   "煤粉仓温度高报警" AT %Q5.1 : Bool;
   "回转窑助燃罗茨风机启动" AT %Q4.7 : Bool;
   "Q3_7" AT %Q3.7 : Bool;
   "Q3_6" AT %Q3.6 : Bool;
   "Q3_5" AT %Q3.5 : Bool;
   "Q3_4" AT %Q3.4 : Bool;
   "Q3_3" AT %Q3.3 : Bool;
   "Q3_2" AT %Q3.2 : Bool;
   "Q3_1" AT %Q3.1 : Bool;
   "Q3_0" AT %Q3.0 : Bool;
   "Q2_7" AT %Q2.7 : Bool;
   "Q2_6" AT %Q2.6 : Bool;
   "Q2_5" AT %Q2.5 : Bool;
   "Q2_4" AT %Q2.4 : Bool;
   "Q2_3" AT %Q2.3 : Bool;
   "Q2_2" AT %Q2.2 : Bool;
   "Q2_1" AT %Q2.1 : Bool;
   "Q2_0" AT %Q2.0 : Bool;
   "Q1_7" AT %Q1.7 : Bool;
   "Q1_1" AT %Q1.1 : Bool;
   "窑尾罩温度输出" AT %QW286 : Int;
   "PQW278" AT %QW278 : Int;
   "4#回转窑富氧调节阀给定" AT %QW276 : Int;
   "助燃罗茨风机频率给定" AT %QW274 : Int;
   "PQW270" AT %QW270 : Int;
   "PQW268" AT %QW268 : Int;
   "PQW266" AT %QW266 : Int;
   "PQW264" AT %QW264 : Int;
   "PQW262" AT %QW262 : Int;
   "PQW260" AT %QW260 : Int;
   "7#配料皮带启动" AT %Q6.6 : Bool;
   "7#配料流量给定" AT %QW300 : Int;
   "6#配料皮带启动" AT %Q6.5 : Bool;
   "6#配料流量给定" AT %QW298 : Int;
   "5#配料皮带启动" AT %Q6.4 : Bool;
   "5#配料流量给定" AT %QW296 : Int;
   "4#配料皮带启动" AT %Q6.3 : Bool;
   "4#配料流量给定" AT %QW294 : Int;
   "3#配料皮带启动" AT %Q6.2 : Bool;
   "3#配料流量给定" AT %QW292 : Int;
   "2#配料皮带启动" AT %Q6.1 : Bool;
   "2#配料流量给定" AT %QW290 : Int;
   "1#配料皮带启动" AT %Q6.0 : Bool;
   "1#配料流量给定" AT %QW288 : Int;
   "闸阀下限" AT %M80.7 : Bool;
   "闸阀上限" AT %M80.6 : Bool;
   "窑体行程下下限停窑计时" AT %M8.1 : Bool;
   "窑体行程上上限停窑计时" AT %M8.0 : Bool;
   "挡轮油站重故障_BOOL" AT %M10.2 : Bool;
   "回转窑转子秤连锁" AT %M80.2 : Bool;
   "从机稀油重故障_BOOL" AT %M10.1 : Bool;
   "从机稀油油差下限停窑计时" AT %M0.3 : Bool;
   "主机稀油重故障_BOOL" AT %M10.0 : Bool;
   "主机稀油油位上限停窑计时" AT %M0.4 : Bool;
   "Tag_4" AT %M1.0 : Bool;
   "Tag_3" AT %M1.1 : Bool;
   "Tag_23" AT %MW74 : Word;
   "Tag_22" AT %MD338 : DWord;
   "Tag_21" AT %MW72 : Word;
   "Tag_20" AT %MD336 : DWord;
   "Tag_2" AT %MW6 : Word;
   "Tag_19" AT %MW68 : Word;
   "Tag_18" AT %MD328 : DWord;
   "Tag_17" AT %M0.0 : Bool;
   "Tag_16" AT %MW62 : Word;
   "Tag_15" AT %M0.1 : Bool;
   "Tag_14" AT %M101.6 : Bool;
   "Tag_12" AT %M101.7 : Bool;
   "Tag_11" AT %MW60 : Word;
   "Tag_1" AT %MW4 : Word;
   "Zhongjianzhi4-1" AT %MD100 : Real;
   "Zhongjianzhi4-2" AT %MD104 : Real;
   "Zhongjianzhi4-3" AT %MD108 : Real;
   "Zhongjianzhi4-4" AT %MD112 : Real;
   "Zhongjianzhi5-1" AT %MD116 : Real;
   "Zhongjianzhi5-2" AT %MD120 : Real;
   "Zhongjianzhi5-3" AT %MD124 : Real;
   "Zhongjianzhi5-4" AT %MD128 : Real;
   "Zhongjianzhi6-1" AT %MD132 : Real;
   "Zhongjianzhi6-2" AT %MD136 : Real;
   "Zhongjianzhi6-3" AT %MD140 : Real;
   "Zhongjianzhi6-4" AT %MD144 : Real;
   "Zhongjianzhi7-1" AT %MD148 : Real;
   "Zhongjianzhi7-2" AT %MD152 : Real;
   "Zhongjianzhi7-3" AT %MD156 : Real;
   "Zhongjianzhi7-4" AT %MD160 : Real;
   "Tag_5" AT %M11.0 : Bool;
   "煤粉仓温度高报警中间量" AT %M102.0 : Bool;
   "煤粉仓温度高报警试验按钮" AT %M102.1 : Bool;
   "提升皮带机打滑故障" AT %M9.0 : Bool;
   "提升皮带机打滑故障复位" AT %M9.1 : Bool;
   "24# 煤粉仓消防阀开阀按钮" AT %M9.2 : Bool;
   "24# 煤粉仓消防阀关阀按钮" AT %M9.3 : Bool;
   "挡轮站启动时间" AT %T10 : Timer;
   "挡轮站停止时间" AT %T11 : Timer;
   "挡轮油站重故障判断时间" AT %T22 : Timer;
   "从稀油站启动时间" AT %T14 : Timer;
   "从稀油站停止时间" AT %T15 : Timer;
   "从机稀油重故障判断时间" AT %T21 : Timer;
   "主稀油站启动时间" AT %T12 : Timer;
   "主稀油站停止时间" AT %T13 : Timer;
   "主机稀油重故障判断时间" AT %T20 : Timer;
   "Tag_9" AT %T112 : Timer;
   "Tag_8" AT %T108 : Timer;
   "Tag_7" AT %T107 : Timer;
   "Tag_35" AT %T38 : Timer;
   "Tag_34" AT %T37 : Timer;
   "Tag_33" AT %T36 : Timer;
   "Tag_32" AT %T35 : Timer;
   "Tag_31" AT %T34 : Timer;
   "Tag_30" AT %T33 : Timer;
   "Tag_29" AT %T32 : Timer;
   "Tag_28" AT %T31 : Timer;
   "Tag_27" AT %T30 : Timer;
   "Tag_25" AT %T101 : Timer;
   "Tag_24" AT %T100 : Timer;
   "Tag_10" AT %T111 : Timer;
   "Tag_6" AT %T113 : Timer;
   "Tag_36" AT %T114 : Timer;
   "Tag_13" AT %C1 : Counter;
   "4#回转窑富氧流量" AT %IW356 : Int;
   "4#回转窑富氧调节阀反馈" AT %IW358 : Int;
   "4#回转窑富氧快切阀开按钮" AT %M9.4 : Bool;
   "4#回转窑富氧快切阀关按钮" AT %M9.5 : Bool;
   "4#回转窑富氧压力" AT %IW354 : Int;
   "4#回转窑富氧压力连锁点" AT %M9.6 : Bool;
   "4#回转窑富氧含量" AT %IW352 : Int;
   "Tag_37" AT %T115 : Timer;
   "4#回转窑富氧连锁投入与解除" AT %M9.7 : Bool;
END_VAR

DATA_BLOCK "DB块"   // DB1
{ S7_Optimized_Access := 'FALSE' }
VERSION : 0.1
   VAR
      STAT0 : Bool;
      STAT1 : Bool;
      STAT2 : Bool;
      STAT3_1 : Bool;
      STAT4_1 : Bool;
      STAT4_2 : Bool;
      "4#回转窑烟气管道闸板上限给定" : Real := 180.0;
      "4#回转窑烟气管道闸板下限给定" : Real := 5.0;
      定量给煤机班累计清零 : Bool;
      定量给煤机日累计清零 : Bool;
      定量给煤机总累计清零 : Bool;
   END_VAR
BEGIN
END_DATA_BLOCK

DATA_BLOCK "DB2_配料站清零按钮"   // DB2
{ S7_Optimized_Access := 'FALSE' }
VERSION : 0.1
   VAR
      "班01-1" : Bool;
      "班01-2" : Bool;
      "班01-3" : Bool;
      "班01-4" : Bool;
      "班01-5" : Bool;
      "班01-6" : Bool;
      "班01-7" : Bool;
      "班01-8" : Bool;
      "日01-1" : Bool;
      "日01-2" : Bool;
      "日01-3" : Bool;
      "日01-4" : Bool;
      "日01-5" : Bool;
      "日01-6" : Bool;
      "日01-7" : Bool;
      "日01-8" : Bool;
      "月01-1" : Bool;
      "月01-2" : Bool;
      "月01-3" : Bool;
      "月01-4" : Bool;
      "月01-5" : Bool;
      "月01-6" : Bool;
      "月01-7" : Bool;
      "月01-8" : Bool;
      "总01-1" : Bool;
      "总01-2" : Bool;
      "总01-3" : Bool;
      "总01-4" : Bool;
      "总01-5" : Bool;
      "总01-6" : Bool;
      "总01-7" : Bool;
      "总01-8" : Bool;
      备用1 : Bool;
      备用2 : Bool;
      备用3 : Bool;
      备用4 : Bool;
      备用5 : Bool;
      备用6 : Bool;
      备用7 : Bool;
      备用8 : Bool;
      备用9 : Bool;
      备用10 : Bool;
      备用11 : Bool;
      备用12 : Bool;
      备用13 : Bool;
      备用14 : Bool;
      备用15 : Bool;
      备用16 : Bool;
   END_VAR
BEGIN
END_DATA_BLOCK

DATA_BLOCK "给煤机班累计DB块"   // DB3
{ S7_Optimized_Access := 'FALSE' }
VERSION : 0.0
// stored: InstanceOfName 累计功能块
"累计功能块"
BEGIN
END_DATA_BLOCK

DATA_BLOCK "给煤机日累计DB块"   // DB4
{ S7_Optimized_Access := 'FALSE' }
VERSION : 0.0
// stored: InstanceOfName 累计功能块
"累计功能块"
BEGIN
END_DATA_BLOCK

DATA_BLOCK "给煤机总累计DB块"   // DB5
{ S7_Optimized_Access := 'FALSE' }
VERSION : 0.0
// stored: InstanceOfName 累计功能块
"累计功能块"
BEGIN
END_DATA_BLOCK

DATA_BLOCK "DB6_皮带秤粘料"   // DB6
{ S7_Optimized_Access := 'FALSE' }
VERSION : 0.1
   VAR
      转子秤给定反馈差值 : Real;
      转子秤给定反馈差值绝对值 : Real;
      real3 : Real;
      real4 : Real;
      real5 : Real;
      real6 : Real;
      real7 : Real;
      real8 : Real;
      real9 : Real;
      real10 : Real;
      real11 : Real;
      real12 : Real;
      real13 : Real;
      real14 : Real;
      real15 : Real;
      real16 : Real;
      real17 : Real;
      real18 : Real;
      real19 : Real;
      real20 : Real;
      转子秤粘料报警 : Bool;
      板式给料机粘料报警 : Bool;
      "1#配料皮带粘料报警" : Bool;
      "2#配料皮带粘料报警" : Bool;
      "3#配料皮带粘料报警" : Bool;
      "4#配料皮带粘料报警" : Bool;
      "5#配料皮带粘料报警" : Bool;
      "6#配料皮带粘料报警" : Bool;
      "7#配料皮带粘料报警" : Bool;
      bool10 : Bool;
      bool11 : Bool;
      bool12 : Bool;
      bool13 : Bool;
      bool14 : Bool;
      bool15 : Bool;
      bool16 : Bool;
      bool17 : Bool;
      bool18 : Bool;
      bool19 : Bool;
      bool20 : Bool;
      bool21 : Bool;
   END_VAR
BEGIN
END_DATA_BLOCK

DATA_BLOCK "DB10"   // DB10
{ S7_Optimized_Access := 'FALSE' }
VERSION : 0.1
   VAR
      "4#回转窑主传转速" : Real := 912.7778;
      "4#回转窑主传电流" : Real := 87.62963;
      "4#回转窑主传转速给定" : Real := 900.0;
      STAT3 : Real;
      "4#回转窑从传转速" : Real := 914.1666;
      "4#回转窑从传电流" : Real := 104.8889;
      STAT6 : Real;
      STAT7 : Real;
      "4#回转窑窑体温度1" : Real := 576.4178;
      "4#回转窑窑体温度2" : Real := 557.3206;
      "4#回转窑窑体温度3" : Real := 803.6747;
      "4#回转窑窑体温度4" : Real := 259.4039;
      "4#回转窑窑体温度5" : Real := 212.934;
      "4#回转窑窑体温度6" : Real := 179.8322;
      STAT14 : Real;
      STAT15 : Real;
      STAT16 : Real;
      STAT17 : Real;
      STAT18 : Real;
      STAT19 : Real;
      "4#回转窑窑尾温度" : Real := 250.1447;
      STAT21 : Real;
      "4#回转窑窑尾负压" : Real := -261.8055;
      STAT23 : Real;
      "4#回转窑煤粉仓温度1" : Real := 35.01157;
      "4#回转窑煤粉仓温度2" : Real := 31.85764;
      "4#回转窑煤粉仓温度3" : Real := 31.97338;
      "4#回转窑煤粉仓温度4" : Real := 35.59028;
      "4#回转窑煤粉仓温度5" : Real := 33.01505;
      "4#回转窑煤粉仓温度6" : Real := 62.41319;
      STAT30 : Real;
      STAT31 : Real;
      STAT32 : Real;
      "4#回转窑助燃罗茨风机运行频率" : Real;
      "4#回转窑助燃罗茨风机运行电流" : Real;
      "4#回转窑助燃罗茨风机频率给定" : Real;
      "4#回转窑转子秤流量" : Real := 3.599826;
      "4#回转窑转子秤流量给定" : Real := 1.0;
      "4#回转窑煤粉仓称重" : Real := 7.06;   // 4#回转窑煤粉仓称重
      STAT39 : Real;
      "4#回转窑送煤风机管道压力" : Real := 10.36458;
      STAT41 : Real;
      "4#回转窑煤粉仓压力" : Real := -3197.917;
      STAT43 : Real;
      "4#回转窑窑头温度" : Real := 208.3333;
      STAT45 : Real;
      "4#回转窑窑头负压" : Real := -120.3125;
      STAT47 : Real;
      "4#回转窑中间仓称重" : Real := 3.21;   // 4#回转窑中间仓称重
      STAT49 : Real;
      "4#回转窑送风风机管道压力" : Real := 10.78125;
      "4#回转窑一次风机频率给定" : Real := 39.0;
      "4#回转窑一次风机运行频率" : Real := 38.80209;
      "4#回转窑二次风机运行频率" : Real := 27.70544;
      "4#回转窑二次风机频率给定" : Real := 28.0;
      STAT55 : Real;
      "4#回转窑一次风机运行电流" : Real := 49.0162;
      "4#回转窑二次风机运行电流" : Real := 57.40625;
      STAT58 : Real;
      STAT59 : Real;
      "4#回转窑支撑挡轮温度A1" : Real := 35.0;
      "4#回转窑支撑挡轮温度A2" : Real := 34.0;
      "4#回转窑支撑挡轮温度A3" : Real := 36.0;
      "4#回转窑支撑挡轮温度A4" : Real := 34.0;
      "4#回转窑支撑挡轮温度B1" : Real := 37.0;
      "4#回转窑支撑挡轮温度B2" : Real := 35.0;
      "4#回转窑支撑挡轮温度B3" : Real := 37.0;
      "4#回转窑支撑挡轮温度B4" : Real := 32.0;
      "4#回转窑支撑挡轮温度C1" : Real := 34.0;
      "4#回转窑支撑挡轮温度C2" : Real := 34.0;
      "4#回转窑支撑挡轮温度C3" : Real := 37.0;
      "4#回转窑支撑挡轮温度C4" : Real := 36.0;
      "4#回转窑支撑挡轮温度D1" : Real := 37.0;
      "4#回转窑支撑挡轮温度D2" : Real := 32.0;
      "4#回转窑支撑挡轮温度D3" : Real := 35.0;
      "4#回转窑支撑挡轮温度D4" : Real := 33.0;
      "4#回转窑支撑挡轮轴温度A1" : Real := 34.0;
      "4#回转窑支撑挡轮轴温度A2" : Real := 34.0;
      "4#回转窑支撑挡轮轴温度A3" : Real := 34.0;
      "4#回转窑支撑挡轮轴温度A4" : Real := 35.0;
      "4#回转窑支撑挡轮轴温度B1" : Real := 32.0;
      "4#回转窑支撑挡轮轴温度B2" : Real := 33.0;
      "4#回转窑支撑挡轮轴温度B3" : Real := 35.0;
      "4#回转窑支撑挡轮轴温度B4" : Real := 34.0;
      "4#回转窑支撑挡轮轴温度C1" : Real := 33.0;
      "4#回转窑支撑挡轮轴温度C2" : Real := 31.0;
      "4#回转窑支撑挡轮轴温度C3" : Real := 35.0;
      "4#回转窑支撑挡轮轴温度C4" : Real := 36.0;
      "4#回转窑支撑挡轮轴温度D1" : Real := 32.0;
      "4#回转窑支撑挡轮轴温度D2" : Real := 35.0;
      "4#回转窑支撑挡轮轴温度D3" : Real := 33.0;
      "4#回转窑支撑挡轮轴温度D4" : Real := 37.0;
      "4#回转窑备用一次风机运行频率" : Real := 0.2170139;
      "4#回转窑备用一次风机频率给定" : Real := 5.0;
      STAT94 : Real;
      "4#回转窑备用一次风机运行电流" : Real := 0.2430556;
      STAT96 : Real;
      STAT97 : Real;
      "4#回转窑窑尾烟气管道标尺高度" : Real := 80.20834;
      "4#回转窑定量给煤机班累计" : Real := 3090.047;
      "4#回转窑定量给煤机日累计" : Real := 3090.047;
      "4#回转窑定量给煤机总累计" : Real := 3090.047;
   END_VAR
BEGIN
END_DATA_BLOCK

DATA_BLOCK "DB12"   // DB12
{ S7_Optimized_Access := 'FALSE' }
VERSION : 0.1
   VAR
      "4#回转窑主传接触器合闸" : Bool;
      "4#回转窑主传接触器分闸" : Bool;
      "4#回转窑主传变频器启动" : Bool;
      "4#回转窑主传变频器停止" : Bool;
      "4#回转窑主机稀油站启动" : Bool;
      "4#回转窑主机稀油站停止" : Bool;
      "4#回转窑从机稀油站启动" : Bool;
      "4#回转窑从机稀油站停止" : Bool;
      STAT8 : Bool;
      STAT9 : Bool;
      STAT10 : Bool;
      STAT11 : Bool;
      STAT12 : Bool;
      STAT13 : Bool;
      STAT14 : Bool;
      STAT15 : Bool;
      "4#回转窑煤粉仓收尘风机启动" : Bool;
      "4#回转窑煤粉仓收尘风机停止" : Bool;
      "4#回转窑转子秤启动" : Bool;
      "4#回转窑转子秤停止" : Bool;
      STAT20 : Bool;
      STAT21 : Bool;
      STAT22 : Bool;
      STAT23 : Bool;
      "4#回转窑窑头护板风机启动" : Bool;
      "4#回转窑窑头护板风机停止" : Bool;
      STAT26 : Bool;
      STAT27 : Bool;
      STAT28 : Bool;
      STAT29 : Bool;
      STAT30 : Bool;
      STAT31 : Bool;
      STAT32 : Bool;
      STAT33 : Bool;
      "4#回转窑干矿提升皮带启动" : Bool;
      "4#回转窑干矿提升皮带停止" : Bool;
      STAT36 : Bool;
      STAT37 : Bool;
      "4#回转窑干矿进料皮带启动" : Bool;
      "4#回转窑干矿进料皮带停止" : Bool;
      STAT40 : Bool;
      STAT41 : Bool;
      STAT42 : Bool;
      STAT43 : Bool;
      STAT44 : Bool;
      STAT45 : Bool;
      "4#回转窑一次风机启动" : Bool;
      "4#回转窑一次风机停止" : Bool;
      "4#回转窑二次风机启动" : Bool;
      "4#回转窑二次风机停止" : Bool;
      STAT50 : Bool;
      STAT51 : Bool;
      STAT52 : Bool;
      STAT53 : Bool;
      "4#回转窑备用一次风机启动" : Bool;
      "4#回转窑备用一次风机停止" : Bool;
      "4#回转窑助燃罗茨风机启动" : Bool;
      "4#回转窑助燃罗茨风机停止" : Bool;
      STAT58 : Bool;
      STAT59 : Bool;
      "4#回转窑挡轮油站启动" : Bool;
      "4#回转窑挡轮油站停止" : Bool;
      STAT62 : Bool;
      STAT63 : Bool;
      "4#回转窑联锁解锁状态" : Bool := TRUE;
      STAT65 : Bool;
      "4#回转窑烟气管道闸板上升" : Bool;
      "4#回转窑烟气管道闸板下降" : Bool;
      STAT68 : Bool;
      STAT69 : Bool;
   END_VAR
BEGIN
END_DATA_BLOCK

DATA_BLOCK "DB20"   // DB20
{ S7_Optimized_Access := 'FALSE' }
VERSION : 0.1
   VAR
      STAT0 : Real := 0.004340278;
      STAT1 : Real := 1.458333;
      STAT2 : Real := 1.252893;
      STAT3 : Real := 33.17708;
      STAT4 : Real := 35.70313;
      STAT5 : Real := 11.45833;
      STAT6 : Real;
      STAT7 : Real;
      STAT8 : Real;
      STAT9 : Real;
      STAT10 : Real;
      STAT11 : Real;
      STAT12 : Real;
      STAT13 : Real;
      STAT14 : Real := 93.51852;
      STAT15 : Real;
      STAT16 : Real;
      STAT17 : Real := 1.44;
      STAT18 : Real := 1.28;
      STAT19 : Real := 32.0;
      STAT20 : Real := 36.0;
      STAT21 : Real := 12.0;
      STAT22 : Real;
      STAT23 : Real;
      STAT24 : Real;
      STAT25 : Real;
      STAT26 : Real;
      STAT27 : Real;
      STAT28 : Real;
      STAT29 : Real;
      STAT30 : Real := 100.0;
      STAT31 : Real;
      STAT32 : Real;
      STAT33 : Real;
      STAT34 : Real := 462.819;
      STAT35 : Real := 462.819;
      STAT36 : Real := 0.9000001;
      STAT37 : Real := 11.40001;
      STAT38 : Real := 2151.148;
      STAT39 : Real := 2151.148;
      STAT40 : Real := 0.8000001;
      STAT41 : Real := 11.30001;
      STAT42 : Real := 1006.201;
      STAT43 : Real := 1006.201;
      STAT44 : Real := 21.0;
      STAT45 : Real := 298.0;
      STAT46 : Real := 14706.0;
      STAT47 : Real := 14706.0;
      STAT48 : Real := 24.0;
      STAT49 : Real := 264.0;
      STAT50 : Real := 22921.0;
      STAT51 : Real := 22921.0;
      STAT52 : Real := 8.0;
      STAT53 : Real := 105.0;
      STAT54 : Real := 26878.0;
      STAT55 : Real := 26878.0;
      STAT56 : Real;
      STAT57 : Real;
      STAT58 : Real := 25069.0;
      STAT59 : Real := 25069.0;
      STAT60 : Real;
      STAT61 : Real;
      STAT62 : Real;
      STAT63 : Real;
      STAT64 : Real;
      STAT65 : Real;
      STAT66 : Real;
      STAT67 : Real;
      STAT68 : Real;
      STAT69 : Real;
      STAT70 : Real;
      STAT71 : Real;
      STAT72 : Real;
      STAT73 : Real;
      STAT74 : Real;
      STAT75 : Real;
      STAT76 : Real;
      STAT77 : Real;
      STAT78 : Real;
      STAT79 : Real;
      STAT80 : Real;
      STAT81 : Real;
      STAT82 : Real;
      STAT83 : Real;
      STAT84 : Real;
      STAT85 : Real;
      STAT86 : Real;
      STAT87 : Real;
      STAT88 : Real := 38.0;
      STAT89 : Real := 28163.0;
      STAT90 : Real := 28163.0;
      STAT91 : Real := 28163.0;
      STAT92 : Bool;
      STAT93 : Bool;
      STAT94 : Bool;
      STAT95 : Bool;
      STAT96 : Bool;
      STAT97 : Bool;
      STAT98 : Bool;
      STAT99 : Bool;
      STAT100 : Bool;
      STAT101 : Bool;
      STAT102 : Bool;
      STAT103 : Bool;
      STAT104 : Bool;
      STAT105 : Bool;
      STAT106 : Bool;
      STAT107 : Bool;
      STAT108 : Bool;
      STAT109 : Bool;
      STAT110 : Bool;
      STAT111 : Bool;
   END_VAR
BEGIN
END_DATA_BLOCK

DATA_BLOCK "DB22"   // DB22
{ S7_Optimized_Access := 'FALSE' }
VERSION : 0.1
   VAR
      STAT0 : Real := 43.89034;
      STAT1 : Real := 38.65741;
      STAT2 : Real := 38.0;
      STAT3 : Bool;
      STAT4 : Bool;
      STAT5 : Bool;
      STAT6 : Bool;
      STAT7 : Bool;
      STAT8 : Bool;
      STAT9 : Bool;
      STAT10 : Bool;
   END_VAR
BEGIN
END_DATA_BLOCK

DATA_BLOCK "数据块_电机温度"   // DB23
{ S7_Optimized_Access := 'FALSE' }
VERSION : 0.1
   VAR
      主电机定子温度 : Real;
      主电机前轴温度 : Real;
      主电机后轴温度 : Real;
      从电机定子温度 : Real;
      从电机前轴温度 : Real;
      从电机后轴温度 : Real;
      "4#回转窑富氧流量" : Real;
      "4#回转窑富氧调节阀反馈" : Real;
      "4#回转窑富氧调节阀给定" : Real;
      "4#回转窑富氧压力" : Real;
      "4#回转窑富氧压力设定" : Real;
      "4#回转窑富氧含量" : Real;
   END_VAR
BEGIN
END_DATA_BLOCK

DATA_BLOCK "DB201"   // DB201
{ S7_Optimized_Access := 'FALSE' }
VERSION : 0.0
// stored: InstanceOfName 给料电机启动块
"给料电机启动块"
BEGIN
END_DATA_BLOCK

DATA_BLOCK "DB202"   // DB202
{ S7_Optimized_Access := 'FALSE' }
VERSION : 0.0
// stored: InstanceOfName 给料电机启动块
"给料电机启动块"
BEGIN
END_DATA_BLOCK

DATA_BLOCK "DB203"   // DB203
{ S7_Optimized_Access := 'FALSE' }
VERSION : 0.0
// stored: InstanceOfName 给料电机启动块
"给料电机启动块"
BEGIN
END_DATA_BLOCK

DATA_BLOCK "DB204"   // DB204
{ S7_Optimized_Access := 'FALSE' }
VERSION : 0.0
// stored: InstanceOfName 给料电机启动块
"给料电机启动块"
BEGIN
END_DATA_BLOCK

DATA_BLOCK "DB205"   // DB205
{ S7_Optimized_Access := 'FALSE' }
VERSION : 0.0
// stored: InstanceOfName 给料电机启动块
"给料电机启动块"
BEGIN
END_DATA_BLOCK

DATA_BLOCK "DB206"   // DB206
{ S7_Optimized_Access := 'FALSE' }
VERSION : 0.0
// stored: InstanceOfName 给料电机启动块
"给料电机启动块"
BEGIN
END_DATA_BLOCK

DATA_BLOCK "DB207"   // DB207
{ S7_Optimized_Access := 'FALSE' }
VERSION : 0.0
// stored: InstanceOfName 给料电机启动块
"给料电机启动块"
BEGIN
END_DATA_BLOCK

DATA_BLOCK "DB208"   // DB208
{ S7_Optimized_Access := 'FALSE' }
VERSION : 0.0
// stored: InstanceOfName 给料电机启动块
"给料电机启动块"
BEGIN
END_DATA_BLOCK

DATA_BLOCK "DB210"   // DB210
{ S7_Optimized_Access := 'FALSE' }
VERSION : 0.0
// stored: InstanceOfName FB11
"FB11"
BEGIN
END_DATA_BLOCK

DATA_BLOCK "DB211"   // DB211
{ S7_Optimized_Access := 'FALSE' }
VERSION : 0.0
// stored: InstanceOfName FB11
"FB11"
BEGIN
END_DATA_BLOCK

DATA_BLOCK "DB212"   // DB212
{ S7_Optimized_Access := 'FALSE' }
VERSION : 0.0
// stored: InstanceOfName FB11
"FB11"
BEGIN
END_DATA_BLOCK

DATA_BLOCK "DB213"   // DB213
{ S7_Optimized_Access := 'FALSE' }
VERSION : 0.1
// stored: InstanceOfName FB11
"FB11"
BEGIN
END_DATA_BLOCK

DATA_BLOCK "DB214"   // DB214
{ S7_Optimized_Access := 'FALSE' }
VERSION : 0.1
// stored: InstanceOfName FB11
"FB11"
BEGIN
END_DATA_BLOCK

DATA_BLOCK "DB215"   // DB215
{ S7_Optimized_Access := 'FALSE' }
VERSION : 0.1
// stored: InstanceOfName FB11
"FB11"
BEGIN
END_DATA_BLOCK

DATA_BLOCK "DB216"   // DB216
{ S7_Optimized_Access := 'FALSE' }
VERSION : 0.1
// stored: InstanceOfName FB11
"FB11"
BEGIN
END_DATA_BLOCK

DATA_BLOCK "DB217"   // DB217
{ S7_Optimized_Access := 'FALSE' }
VERSION : 0.0
// stored: InstanceOfName FB9
"FB9"
BEGIN
END_DATA_BLOCK

DATA_BLOCK "DB218"   // DB218
{ S7_Optimized_Access := 'FALSE' }
VERSION : 0.1
// stored: InstanceOfName FB9
"FB9"
BEGIN
END_DATA_BLOCK

DATA_BLOCK "DB219"   // DB219
{ S7_Optimized_Access := 'FALSE' }
VERSION : 0.1
// stored: InstanceOfName FB9
"FB9"
BEGIN
END_DATA_BLOCK

DATA_BLOCK "DB220"   // DB220
{ S7_Optimized_Access := 'FALSE' }
VERSION : 0.0
// stored: InstanceOfName FB11
"FB11"
BEGIN
END_DATA_BLOCK

DATA_BLOCK "DB221"   // DB221
{ S7_Optimized_Access := 'FALSE' }
VERSION : 0.0
// stored: InstanceOfName FB11
"FB11"
BEGIN
END_DATA_BLOCK

DATA_BLOCK "DB222"   // DB222
{ S7_Optimized_Access := 'FALSE' }
VERSION : 0.0
// stored: InstanceOfName FB11
"FB11"
BEGIN
END_DATA_BLOCK

DATA_BLOCK "DB223"   // DB223
{ S7_Optimized_Access := 'FALSE' }
VERSION : 0.1
// stored: InstanceOfName FB9
"FB9"
BEGIN
END_DATA_BLOCK

DATA_BLOCK "DB224"   // DB224
{ S7_Optimized_Access := 'FALSE' }
VERSION : 0.1
// stored: InstanceOfName FB9
"FB9"
BEGIN
END_DATA_BLOCK

FUNCTION_BLOCK "给料电机启动块"   // FB8, LAD
{ S7_Optimized_Access := 'FALSE' }
VERSION : 0.1
   VAR_INPUT
      IN0 : Bool;
      IN1 : Bool;
      IN2 : Bool;
      IN3 : Bool;
      IN4 : Bool;
      IN5 : Bool;
   END_VAR
   VAR_IN_OUT
      OUT6 : Bool;
   END_VAR
BEGIN

REGION Network 1
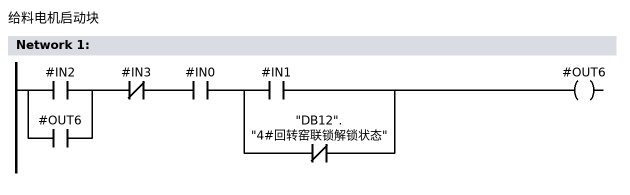
   RUNG wire#powerrail
      Contact( #IN2 )
      wire#w1
      I_Contact( #IN3 )
      Contact( #IN0 )
      wire#w2
      Contact( #IN1 )
      wire#w3
      Coil( #OUT6 )
   END_RUNG
   RUNG wire#powerrail
      Contact( #OUT6 )
   END_RUNG wire#w1
   RUNG wire#w2
      I_Contact( "DB12"."4#回转窑联锁解锁状态" )
   END_RUNG wire#w3
   // the same network as SCL:
   #OUT6 := (#IN2 OR #OUT6) AND NOT #IN3 AND #IN0 AND (#IN1 OR NOT "DB12"."4#回转窑联锁解锁状态");
END_REGION

REGION Network 2 (STL)
         SET;
         SAVE;
END_REGION
END_FUNCTION_BLOCK

FUNCTION_BLOCK "FB9"   // FB9, LAD
{ S7_Optimized_Access := 'FALSE' }
VERSION : 0.1
   VAR_INPUT
      IN0 : Bool;
      IN1 : Bool;
      IN2 : Bool;
      IN3 : Bool;
      IN4 : Bool;
   END_VAR
   VAR_OUTPUT
      OUT5 : Real;
      OUT6 : Real;
      OUT7 : Real;
      OUT8 : Real;
   END_VAR
   VAR
      STAT9 : Real;
      STAT10 : Real;
      STAT11 : Real;
      STAT12 : Real;
      STAT13 : Bool;
   END_VAR
BEGIN

REGION Network 1
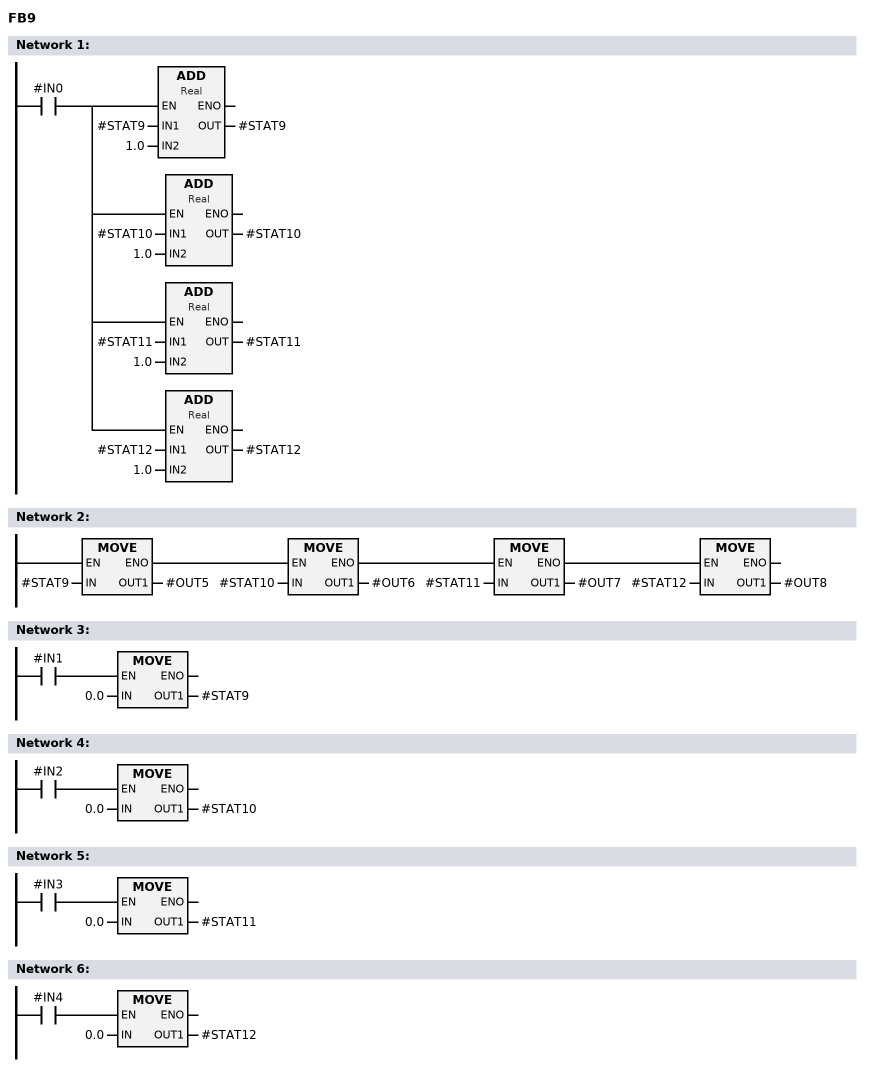
   RUNG wire#powerrail
      Contact( #IN0 )
      wire#w1
      { S7_Templates := "SrcType := Real"; S7_GenerateENO := "TRUE" } Add(in1 := #STAT9, in2 := 1.0, out => #STAT9)
   END_RUNG
   RUNG wire#w1
      { S7_Templates := "SrcType := Real"; S7_GenerateENO := "TRUE" } Add(in1 := #STAT10, in2 := 1.0, out => #STAT10)
   END_RUNG
   RUNG wire#w1
      { S7_Templates := "SrcType := Real"; S7_GenerateENO := "TRUE" } Add(in1 := #STAT11, in2 := 1.0, out => #STAT11)
   END_RUNG
   RUNG wire#w1
      { S7_Templates := "SrcType := Real"; S7_GenerateENO := "TRUE" } Add(in1 := #STAT12, in2 := 1.0, out => #STAT12)
   END_RUNG
   // the same network as SCL:
   IF #IN0 THEN
       #STAT9 := #STAT9 + 1.0;
       #STAT10 := #STAT10 + 1.0;
       #STAT11 := #STAT11 + 1.0;
       #STAT12 := #STAT12 + 1.0;
   END_IF;
END_REGION

REGION Network 2
   RUNG wire#powerrail
      { S7_GenerateENO := "TRUE" } Move(in := #STAT9, out1 => #OUT5)
      { S7_GenerateENO := "TRUE" } Move(in := #STAT10, out1 => #OUT6)
      { S7_GenerateENO := "TRUE" } Move(in := #STAT11, out1 => #OUT7)
      { S7_GenerateENO := "TRUE" } Move(in := #STAT12, out1 => #OUT8)
   END_RUNG
   // the same network as SCL:
   // ENO of a box is taken as its EN; it also drops when the box reports an error
   #OUT5 := #STAT9;
   #OUT6 := #STAT10;
   #OUT7 := #STAT11;
   #OUT8 := #STAT12;
END_REGION

REGION Network 3
   RUNG wire#powerrail
      Contact( #IN1 )
      { S7_GenerateENO := "TRUE" } Move(in := 0.0, out1 => #STAT9)
   END_RUNG
   // the same network as SCL:
   IF #IN1 THEN #STAT9 := 0.0; END_IF;
END_REGION

REGION Network 4
   RUNG wire#powerrail
      Contact( #IN2 )
      { S7_GenerateENO := "TRUE" } Move(in := 0.0, out1 => #STAT10)
   END_RUNG
   // the same network as SCL:
   IF #IN2 THEN #STAT10 := 0.0; END_IF;
END_REGION

REGION Network 5
   RUNG wire#powerrail
      Contact( #IN3 )
      { S7_GenerateENO := "TRUE" } Move(in := 0.0, out1 => #STAT11)
   END_RUNG
   // the same network as SCL:
   IF #IN3 THEN #STAT11 := 0.0; END_IF;
END_REGION

REGION Network 6
   RUNG wire#powerrail
      Contact( #IN4 )
      { S7_GenerateENO := "TRUE" } Move(in := 0.0, out1 => #STAT12)
   END_RUNG
   // the same network as SCL:
   IF #IN4 THEN #STAT12 := 0.0; END_IF;
END_REGION

REGION Network 7 (STL)
         SET;
         SAVE;
END_REGION
END_FUNCTION_BLOCK

FUNCTION_BLOCK "累计功能块"   // FB10, STL
{ S7_Optimized_Access := 'FALSE' }
VERSION : 0.1
   VAR_INPUT
      IN0 : Real;
      IN1 : Bool;
   END_VAR
   VAR_OUTPUT
      OUT2 : Real;
   END_VAR
   VAR
      STAT3 : Real;
      STAT4 : Real;
      STAT5 : Real;
   END_VAR
BEGIN

REGION Network 1
         A(;
         A(;
         A(;
         L     #IN0;
         L     3600.0;
         /R;
         T     #STAT3;
         AN    OV;
         SAVE;
         CLR;
         A     BR;
         );
         JNB   M001;
         L     #STAT3;
         L     10.0;
         /R;
         T     #STAT4;
         AN    OV;
         SAVE;
         CLR;
   M001: A     BR;
         );
         JNB   M002;
         L     #STAT4;
         L     #STAT5;
         +R;
         T     #STAT5;
         AN    OV;
         SAVE;
         CLR;
   M002: A     BR;
         );
         JNB   M003;
         L     #STAT5;
         T     #OUT2;
   M003: NOP   0;
END_REGION

REGION Network 2
         A     #IN1;
         =     %L0.0;
         A     %L0.0;
         JNB   M004;
         L     0.0;
         T     #STAT3;
   M004: NOP   0;
         A     %L0.0;
         JNB   M005;
         L     0.0;
         T     #STAT4;
   M005: NOP   0;
         A     %L0.0;
         JNB   M006;
         L     0.0;
         T     #STAT5;
   M006: NOP   0;
END_REGION

REGION Network 3
         SET;
         SAVE;
END_REGION
END_FUNCTION_BLOCK

FUNCTION_BLOCK "FB11"   // FB11, LAD
{ S7_Optimized_Access := 'FALSE' }
VERSION : 0.1
   VAR_INPUT
      IN0 : Bool;
      IN1 : Bool;
      IN2 : Bool;
      IN3 : Bool;
      IN4 : Bool;
   END_VAR
   VAR_OUTPUT
      OUT5 : Real;
      OUT6 : Real;
      OUT7 : Real;
      OUT8 : Real;
   END_VAR
   VAR
      STAT9 : Real;
      STAT10 : Real;
      STAT11 : Real;
      STAT12 : Real;
      STAT13 : Bool;
   END_VAR
BEGIN

REGION Network 1
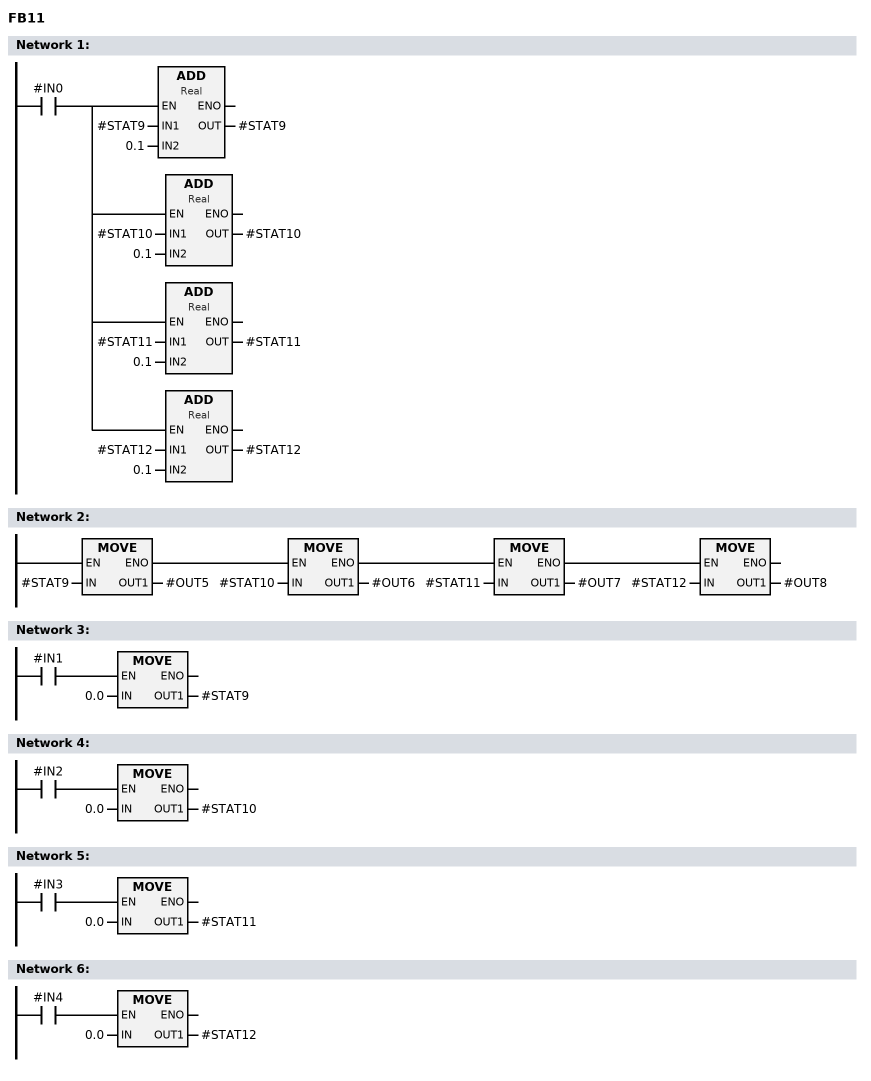
   RUNG wire#powerrail
      Contact( #IN0 )
      wire#w1
      { S7_Templates := "SrcType := Real"; S7_GenerateENO := "TRUE" } Add(in1 := #STAT9, in2 := 0.1, out => #STAT9)
   END_RUNG
   RUNG wire#w1
      { S7_Templates := "SrcType := Real"; S7_GenerateENO := "TRUE" } Add(in1 := #STAT10, in2 := 0.1, out => #STAT10)
   END_RUNG
   RUNG wire#w1
      { S7_Templates := "SrcType := Real"; S7_GenerateENO := "TRUE" } Add(in1 := #STAT11, in2 := 0.1, out => #STAT11)
   END_RUNG
   RUNG wire#w1
      { S7_Templates := "SrcType := Real"; S7_GenerateENO := "TRUE" } Add(in1 := #STAT12, in2 := 0.1, out => #STAT12)
   END_RUNG
   // the same network as SCL:
   IF #IN0 THEN
       #STAT9 := #STAT9 + 0.1;
       #STAT10 := #STAT10 + 0.1;
       #STAT11 := #STAT11 + 0.1;
       #STAT12 := #STAT12 + 0.1;
   END_IF;
END_REGION

REGION Network 2
   RUNG wire#powerrail
      { S7_GenerateENO := "TRUE" } Move(in := #STAT9, out1 => #OUT5)
      { S7_GenerateENO := "TRUE" } Move(in := #STAT10, out1 => #OUT6)
      { S7_GenerateENO := "TRUE" } Move(in := #STAT11, out1 => #OUT7)
      { S7_GenerateENO := "TRUE" } Move(in := #STAT12, out1 => #OUT8)
   END_RUNG
   // the same network as SCL:
   // ENO of a box is taken as its EN; it also drops when the box reports an error
   #OUT5 := #STAT9;
   #OUT6 := #STAT10;
   #OUT7 := #STAT11;
   #OUT8 := #STAT12;
END_REGION

REGION Network 3
   RUNG wire#powerrail
      Contact( #IN1 )
      { S7_GenerateENO := "TRUE" } Move(in := 0.0, out1 => #STAT9)
   END_RUNG
   // the same network as SCL:
   IF #IN1 THEN #STAT9 := 0.0; END_IF;
END_REGION

REGION Network 4
   RUNG wire#powerrail
      Contact( #IN2 )
      { S7_GenerateENO := "TRUE" } Move(in := 0.0, out1 => #STAT10)
   END_RUNG
   // the same network as SCL:
   IF #IN2 THEN #STAT10 := 0.0; END_IF;
END_REGION

REGION Network 5
   RUNG wire#powerrail
      Contact( #IN3 )
      { S7_GenerateENO := "TRUE" } Move(in := 0.0, out1 => #STAT11)
   END_RUNG
   // the same network as SCL:
   IF #IN3 THEN #STAT11 := 0.0; END_IF;
END_REGION

REGION Network 6
   RUNG wire#powerrail
      Contact( #IN4 )
      { S7_GenerateENO := "TRUE" } Move(in := 0.0, out1 => #STAT12)
   END_RUNG
   // the same network as SCL:
   IF #IN4 THEN #STAT12 := 0.0; END_IF;
END_REGION

REGION Network 7 (STL)
         SET;
         SAVE;
END_REGION
END_FUNCTION_BLOCK

FUNCTION "回转窑系统" : Void   // FC1, LAD
{ S7_Optimized_Access := 'FALSE' }
VERSION : 0.1
BEGIN

REGION Network 1
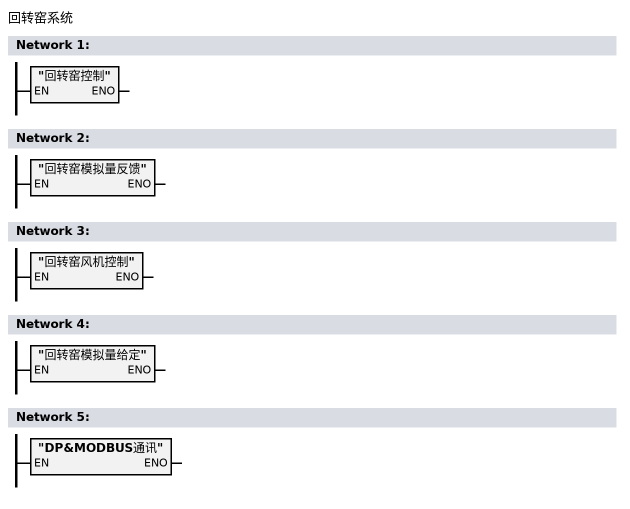
   RUNG wire#powerrail
      "回转窑控制"()
   END_RUNG
   // the same network as SCL:
   "回转窑控制"();
END_REGION

REGION Network 2
   RUNG wire#powerrail
      "回转窑模拟量反馈"()
   END_RUNG
   // the same network as SCL:
   "回转窑模拟量反馈"();
END_REGION

REGION Network 3
   RUNG wire#powerrail
      "回转窑风机控制"()
   END_RUNG
   // the same network as SCL:
   "回转窑风机控制"();
END_REGION

REGION Network 4
   RUNG wire#powerrail
      "回转窑模拟量给定"()
   END_RUNG
   // the same network as SCL:
   "回转窑模拟量给定"();
END_REGION

REGION Network 5
   RUNG wire#powerrail
      "DP&MODBUS通讯"()
   END_RUNG
   // the same network as SCL:
   "DP&MODBUS通讯"();
END_REGION
END_FUNCTION

FUNCTION "配料系统" : Void   // FC2, LAD
{ S7_Optimized_Access := 'FALSE' }
VERSION : 0.1
BEGIN

REGION Network 1
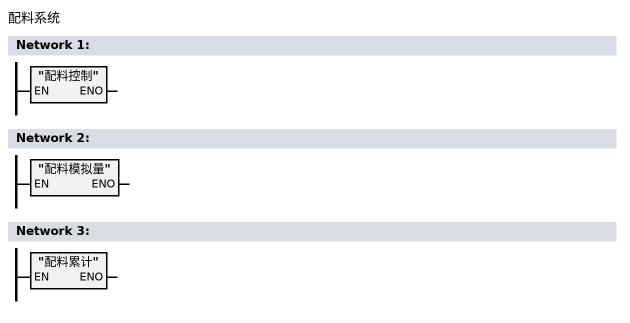
   RUNG wire#powerrail
      "配料控制"()
   END_RUNG
   // the same network as SCL:
   "配料控制"();
END_REGION

REGION Network 2
   RUNG wire#powerrail
      "配料模拟量"()
   END_RUNG
   // the same network as SCL:
   "配料模拟量"();
END_REGION

REGION Network 3
   RUNG wire#powerrail
      "配料累计"()
   END_RUNG
   // the same network as SCL:
   "配料累计"();
END_REGION
END_FUNCTION

FUNCTION "FC4_粘料" : Void   // FC4, LAD
{ S7_Optimized_Access := 'TRUE' }
VERSION : 0.1
   VAR_TEMP   // added for the SCL form of the ladder/FBD networks
      _w1 : Bool;
      _w2 : Bool;
   END_VAR
BEGIN

REGION Network 1